
(*与上位机通讯程序*)
ComConveyor70104(ConveyorIO:= ConveyorIO70140_1,CommunicationIO:= ComConveyorIO70104);
ComConveyor70106(ConveyorIO:= ConveyorIO70140,CommunicationIO:= ComConveyorIO70106);(*线体更改*)
ComConveyor70144(ConveyorIO:= ConveyorIO70144,CommunicationIO:= ComConveyorIO70144);
ComConveyor70152(ConveyorIO:= ConveyorIO70152,CommunicationIO:= ComConveyorIO70152);
ComConveyor70146(ConveyorIO:= ConveyorIO70146,CommunicationIO:= ComConveyorIO70146);
ComConveyor70195(ConveyorIO:= ConveyorIO70195,CommunicationIO:= ComConveyorIO70195);
ComConveyor70147(ConveyorIO:= ConveyorIO70147,CommunicationIO:= ComConveyorIO70147);
ComConveyor70196(ConveyorIO:= ConveyorIO70196,CommunicationIO:= ComConveyorIO70196);
ComConveyor70154(ConveyorIO:= ConveyorIO70154,CommunicationIO:= ComConveyorIO70154);
ComConveyor70199(ConveyorIO:= ConveyorIO70199,CommunicationIO:= ComConveyorIO70199);
ComConveyor70155(ConveyorIO:= ConveyorIO70155,CommunicationIO:= ComConveyorIO70155);
ComConveyor701100(ConveyorIO:= ConveyorIO701100,CommunicationIO:= ComConveyorIO701100);
ComConveyor701115(ConveyorIO:= ConveyorIO701115,CommunicationIO:= ComConveyorIO701115);
ComConveyor701114(ConveyorIO:= ConveyorIO701114,CommunicationIO:= ComConveyorIO701114);
ComConveyor70197(ConveyorIO:= ConveyorIO70197,CommunicationIO:= ComConveyorIO70197);
ComConveyor70150(ConveyorIO:= ConveyorIO70150,CommunicationIO:= ComConveyorIO70150);
ComConveyor70151(ConveyorIO:= ConveyorIO70151,CommunicationIO:= ComConveyorIO70151);
ComConveyor70198(ConveyorIO:= ConveyorIO70198,CommunicationIO:= ComConveyorIO70198);
ComConveyor701101(ConveyorIO:= ConveyorIO701101,CommunicationIO:= ComConveyorIO701101);
ComConveyor70158(ConveyorIO:= ConveyorIO70158,CommunicationIO:= ComConveyorIO70158);
ComConveyor701111(ConveyorIO:= ConveyorIO701111,CommunicationIO:= ComConveyorIO701111);
ComConveyor70148(ConveyorIO:= ConveyorIO70148,CommunicationIO:= ComConveyorIO70148);
ComConveyor70156(ConveyorIO:= ConveyorIO70156,CommunicationIO:= ComConveyorIO70156);
ComConveyor701116(ConveyorIO:= ConveyorIO701116,CommunicationIO:= ComConveyorIO701116);
ComConveyor70164(ConveyorIO:= ConveyorIO70164,CommunicationIO:= ComConveyorIO70164);
ComConveyor70174(ConveyorIO:= ConveyorIO70174,CommunicationIO:= ComConveyorIO70174);
ComConveyor70169(ConveyorIO:= ConveyorIO70169,CommunicationIO:= ComConveyorIO70169);
ComConveyor70170(ConveyorIO:= ConveyorIO70170,CommunicationIO:= ComConveyorIO70170);
ComConveyor70160(ConveyorIO:= ConveyorIO70160,CommunicationIO:= ComConveyorIO70160);
ComConveyor70162(ConveyorIO:= ConveyorIO70162,CommunicationIO:= ComConveyorIO70162);
ComConveyor701103(ConveyorIO:= ConveyorIO701103,CommunicationIO:= ComConveyorIO701103);
ComConveyor70163(ConveyorIO:= ConveyorIO70163,CommunicationIO:= ComConveyorIO70163);
ComConveyor701104(ConveyorIO:= ConveyorIO701104,CommunicationIO:= ComConveyorIO701104);
ComConveyor701102(ConveyorIO:= ConveyorIO701102,CommunicationIO:= ComConveyorIO701102);
ComConveyor70159(ConveyorIO:= ConveyorIO70159,CommunicationIO:= ComConveyorIO70159);
ComConveyor701120(ConveyorIO:= ConveyorIO701120,CommunicationIO:= ComConveyorIO701120);
ComConveyor701119(ConveyorIO:= ConveyorIO701119,CommunicationIO:= ComConveyorIO701119);
(*ComConveyor70111(ConveyorIO:= ConveyorIO70111,CommunicationIO:= ComConveyorIO70111);
ComConveyor70112(ConveyorIO:= ConveyorIO70112,CommunicationIO:= ComConveyorIO70112);
ComConveyor701105(ConveyorIO:= ConveyorIO701105,CommunicationIO:= ComConveyorIO701105);
ComConveyor70113(ConveyorIO:= ConveyorIO70113,CommunicationIO:= ComConveyorIO70113);
ComConveyor701106(ConveyorIO:= ConveyorIO701106,CommunicationIO:= ComConveyorIO701106);
ComConveyor70114(ConveyorIO:= ConveyorIO70114,CommunicationIO:= ComConveyorIO70114);
ComConveyor70116(ConveyorIO:= ConveyorIO70116,CommunicationIO:= ComConveyorIO70116);
ComConveyor70119(ConveyorIO:= ConveyorIO70119,CommunicationIO:= ComConveyorIO70119);
ComConveyor70120(ConveyorIO:= ConveyorIO70120,CommunicationIO:= ComConveyorIO70120);
ComConveyor701107(ConveyorIO:= ConveyorIO701107,CommunicationIO:= ComConveyorIO701107);
ComConveyor70121(ConveyorIO:= ConveyorIO70121,CommunicationIO:= ComConveyorIO70121);
ComConveyor701108(ConveyorIO:= ConveyorIO701108,CommunicationIO:= ComConveyorIO701108);
ComConveyor70122(ConveyorIO:= ConveyorIO70122,CommunicationIO:= ComConveyorIO70122);
ComConveyor70124(ConveyorIO:= ConveyorIO70124,CommunicationIO:= ComConveyorIO70124);
ComConveyor70127(ConveyorIO:= ConveyorIO70127,CommunicationIO:= ComConveyorIO70127);
ComConveyor70128(ConveyorIO:= ConveyorIO70128,CommunicationIO:= ComConveyorIO70128);
ComConveyor701109(ConveyorIO:= ConveyorIO701109,CommunicationIO:= ComConveyorIO701109);
ComConveyor70129(ConveyorIO:= ConveyorIO70129,CommunicationIO:= ComConveyorIO70129);
ComConveyor701110(ConveyorIO:= ConveyorIO701110,CommunicationIO:= ComConveyorIO701110);
ComConveyor70184(ConveyorIO:= ConveyorIO70184,CommunicationIO:= ComConveyorIO70184);*)

ComConveyorIO70104.i_iResponsPCPLC:=D2000; 
ComConveyorIO70104.i_iTypeInfoPCPLC:=D2001;
ComConveyorIO70104.i_iReadWriteFlagPCPLC:=D2005; 
ComConveyorIO70104.i_iTaskProcessFlagPCPLC:=D2006; 
ComConveyorIO70104.i_iCommandPCPLC:=D2007; 
ComConveyorIO70104.i_iTaskIDPCPLC:=D2008; 
DMOV(TRUE,D2009,ComConveyorIO70104.i_diDestinationDevicePCPLC); 
ComConveyorIO70104.i_iProductIDPCPLC:=D2011;
D3000:=ComConveyorIO70104.o_iRequestPLCPC; 
D3001:=ComConveyorIO70104.o_iForceInportPLCPC;
D3002:=ComConveyorIO70104.o_iFolderNumberPLCPC;
D3003:=ComConveyorIO70104.o_iEmptyPLCPC;
D3005:=ComConveyorIO70104.o_iReadWriteFlagPLCPC; 
D3006:=ComConveyorIO70104.o_iDeviceStatusPLCPC; 
D3007:=ComConveyorIO70104.o_iTaskIDPLCPC; 
D3008:=ComConveyorIO70104.o_iProductIDPLCPC;

ComConveyorIO70106.i_iTypeInfoPCPLC:=D2031;
ComConveyorIO70106.i_iReadWriteFlagPCPLC:=D2035; 
ComConveyorIO70106.i_iTaskProcessFlagPCPLC:=D2036; 
ComConveyorIO70106.i_iCommandPCPLC:=D2037; 
ComConveyorIO70106.i_iTaskIDPCPLC:=D2038; 
DMOV(TRUE,D2039,ComConveyorIO70106.i_diDestinationDevicePCPLC); 
ComConveyorIO70106.i_iProductIDPCPLC:=D2041;
D3030:=ComConveyorIO70106.o_iRequestPLCPC; 
D3031:=ComConveyorIO70106.o_iForceInportPLCPC;
D3032:=ComConveyorIO70106.o_iFolderNumberPLCPC;
D3033:=ComConveyorIO70106.o_iEmptyPLCPC;
D3035:=ComConveyorIO70106.o_iReadWriteFlagPLCPC; 
D3036:=ComConveyorIO70106.o_iDeviceStatusPLCPC; 
D3037:=ComConveyorIO70106.o_iTaskIDPLCPC; 
D3038:=ComConveyorIO70106.o_iProductIDPLCPC;
ComConveyorIO70144.i_iResponsPCPLC:=D2045; 
ComConveyorIO70144.i_iTypeInfoPCPLC:=D2046;
ComConveyorIO70144.i_iReadWriteFlagPCPLC:=D2050; 
ComConveyorIO70144.i_iTaskProcessFlagPCPLC:=D2051; 
ComConveyorIO70144.i_iCommandPCPLC:=D2052; 
ComConveyorIO70144.i_iTaskIDPCPLC:=D2053; 
DMOV(TRUE,D2054,ComConveyorIO70144.i_diDestinationDevicePCPLC); 
ComConveyorIO70144.i_iProductIDPCPLC:=D2056;
D3045:=ComConveyorIO70144.o_iRequestPLCPC; 
D3046:=ComConveyorIO70144.o_iForceInportPLCPC;
D3047:=ComConveyorIO70144.o_iFolderNumberPLCPC;
D3048:=ComConveyorIO70144.o_iEmptyPLCPC;
D3050:=ComConveyorIO70144.o_iReadWriteFlagPLCPC; 
D3051:=ComConveyorIO70144.o_iDeviceStatusPLCPC; 
D3052:=ComConveyorIO70144.o_iTaskIDPLCPC; 
D3053:=ComConveyorIO70144.o_iProductIDPLCPC;
ComConveyorIO70152.i_iResponsPCPLC:=D2060; 
ComConveyorIO70152.i_iTypeInfoPCPLC:=D2061;
ComConveyorIO70152.i_iReadWriteFlagPCPLC:=D2065; 
ComConveyorIO70152.i_iTaskProcessFlagPCPLC:=D2066; 
ComConveyorIO70152.i_iCommandPCPLC:=D2067; 
ComConveyorIO70152.i_iTaskIDPCPLC:=D2068; 
DMOV(TRUE,D2069,ComConveyorIO70152.i_diDestinationDevicePCPLC); 
ComConveyorIO70152.i_iProductIDPCPLC:=D2071;
D3060:=ComConveyorIO70152.o_iRequestPLCPC; 
D3061:=ComConveyorIO70152.o_iForceInportPLCPC;
D3062:=ComConveyorIO70152.o_iFolderNumberPLCPC;
D3063:=ComConveyorIO70152.o_iEmptyPLCPC;
D3065:=ComConveyorIO70152.o_iReadWriteFlagPLCPC; 
D3066:=ComConveyorIO70152.o_iDeviceStatusPLCPC; 
D3067:=ComConveyorIO70152.o_iTaskIDPLCPC; 
D3068:=ComConveyorIO70152.o_iProductIDPLCPC;
ComConveyorIO70146.i_iResponsPCPLC:=D2075; 
ComConveyorIO70146.i_iTypeInfoPCPLC:=D2076;
ComConveyorIO70146.i_iReadWriteFlagPCPLC:=D2080; 
ComConveyorIO70146.i_iTaskProcessFlagPCPLC:=D2081; 
ComConveyorIO70146.i_iCommandPCPLC:=D2082; 
ComConveyorIO70146.i_iTaskIDPCPLC:=D2083; 
DMOV(TRUE,D2084,ComConveyorIO70146.i_diDestinationDevicePCPLC); 
ComConveyorIO70146.i_iProductIDPCPLC:=D2086;
D3075:=ComConveyorIO70146.o_iRequestPLCPC; 
D3076:=ComConveyorIO70146.o_iForceInportPLCPC;
D3077:=ComConveyorIO70146.o_iFolderNumberPLCPC;
D3078:=ComConveyorIO70146.o_iEmptyPLCPC;
D3080:=ComConveyorIO70146.o_iReadWriteFlagPLCPC; 
D3081:=ComConveyorIO70146.o_iDeviceStatusPLCPC; 
D3082:=ComConveyorIO70146.o_iTaskIDPLCPC; 
D3083:=ComConveyorIO70146.o_iProductIDPLCPC;
ComConveyorIO70195.i_iResponsPCPLC:=D2090; 
ComConveyorIO70195.i_iTypeInfoPCPLC:=D2091;
ComConveyorIO70195.i_iReadWriteFlagPCPLC:=D2095; 
ComConveyorIO70195.i_iTaskProcessFlagPCPLC:=D2096; 
ComConveyorIO70195.i_iCommandPCPLC:=D2097; 
ComConveyorIO70195.i_iTaskIDPCPLC:=D2098; 
DMOV(TRUE,D2099,ComConveyorIO70195.i_diDestinationDevicePCPLC); 
ComConveyorIO70195.i_iProductIDPCPLC:=D2101;
D3090:=ComConveyorIO70195.o_iRequestPLCPC; 
D3091:=ComConveyorIO70195.o_iForceInportPLCPC;
D3092:=ComConveyorIO70195.o_iFolderNumberPLCPC;
D3093:=ComConveyorIO70195.o_iEmptyPLCPC;
D3095:=ComConveyorIO70195.o_iReadWriteFlagPLCPC; 
D3096:=ComConveyorIO70195.o_iDeviceStatusPLCPC; 
D3097:=ComConveyorIO70195.o_iTaskIDPLCPC; 
D3098:=ComConveyorIO70195.o_iProductIDPLCPC;
ComConveyorIO70147.i_iResponsPCPLC:=D2105; 
ComConveyorIO70147.i_iTypeInfoPCPLC:=D2106;
ComConveyorIO70147.i_iReadWriteFlagPCPLC:=D2110; 
ComConveyorIO70147.i_iTaskProcessFlagPCPLC:=D2111; 
ComConveyorIO70147.i_iCommandPCPLC:=D2112; 
ComConveyorIO70147.i_iTaskIDPCPLC:=D2113; 
DMOV(TRUE,D2114,ComConveyorIO70147.i_diDestinationDevicePCPLC); 
ComConveyorIO70147.i_iProductIDPCPLC:=D2116;
D3105:=ComConveyorIO70147.o_iRequestPLCPC; 
D3106:=ComConveyorIO70147.o_iForceInportPLCPC;
D3107:=ComConveyorIO70147.o_iFolderNumberPLCPC;
D3108:=ComConveyorIO70147.o_iEmptyPLCPC;
D3110:=ComConveyorIO70147.o_iReadWriteFlagPLCPC; 
D3111:=ComConveyorIO70147.o_iDeviceStatusPLCPC; 
D3112:=ComConveyorIO70147.o_iTaskIDPLCPC; 
D3113:=ComConveyorIO70147.o_iProductIDPLCPC;
ComConveyorIO70196.i_iResponsPCPLC:=D2120; 
ComConveyorIO70196.i_iTypeInfoPCPLC:=D2121;
ComConveyorIO70196.i_iReadWriteFlagPCPLC:=D2125; 
ComConveyorIO70196.i_iTaskProcessFlagPCPLC:=D2126; 
ComConveyorIO70196.i_iCommandPCPLC:=D2127; 
ComConveyorIO70196.i_iTaskIDPCPLC:=D2128; 
DMOV(TRUE,D2129,ComConveyorIO70196.i_diDestinationDevicePCPLC); 
ComConveyorIO70196.i_iProductIDPCPLC:=D2131;	
D3120:=ComConveyorIO70196.o_iRequestPLCPC; 
D3121:=ComConveyorIO70196.o_iForceInportPLCPC;
D3122:=ComConveyorIO70196.o_iFolderNumberPLCPC;
D3123:=ComConveyorIO70196.o_iEmptyPLCPC;
D3125:=ComConveyorIO70196.o_iReadWriteFlagPLCPC; 
D3126:=ComConveyorIO70196.o_iDeviceStatusPLCPC; 
D3127:=ComConveyorIO70196.o_iTaskIDPLCPC; 
D3128:=ComConveyorIO70196.o_iProductIDPLCPC;
ComConveyorIO70154.i_iResponsPCPLC:=D2135; 
ComConveyorIO70154.i_iTypeInfoPCPLC:=D2136;
ComConveyorIO70154.i_iReadWriteFlagPCPLC:=D2140; 
ComConveyorIO70154.i_iTaskProcessFlagPCPLC:=D2141; 
ComConveyorIO70154.i_iCommandPCPLC:=D2142; 
ComConveyorIO70154.i_iTaskIDPCPLC:=D2143; 
DMOV(TRUE,D2144,ComConveyorIO70154.i_diDestinationDevicePCPLC); 
ComConveyorIO70154.i_iProductIDPCPLC:=D2146;
D3135:=ComConveyorIO70154.o_iRequestPLCPC; 
D3136:=ComConveyorIO70154.o_iForceInportPLCPC;
D3137:=ComConveyorIO70154.o_iFolderNumberPLCPC;
D3138:=ComConveyorIO70154.o_iEmptyPLCPC;
D3140:=ComConveyorIO70154.o_iReadWriteFlagPLCPC; 
D3141:=ComConveyorIO70154.o_iDeviceStatusPLCPC; 
D3142:=ComConveyorIO70154.o_iTaskIDPLCPC; 
D3143:=ComConveyorIO70154.o_iProductIDPLCPC;
ComConveyorIO70199.i_iResponsPCPLC:=D2150; 
ComConveyorIO70199.i_iTypeInfoPCPLC:=D2151;
ComConveyorIO70199.i_iReadWriteFlagPCPLC:=D2155; 
ComConveyorIO70199.i_iTaskProcessFlagPCPLC:=D2156; 
ComConveyorIO70199.i_iCommandPCPLC:=D2157; 
ComConveyorIO70199.i_iTaskIDPCPLC:=D2158; 
DMOV(TRUE,D2159,ComConveyorIO70199.i_diDestinationDevicePCPLC); 
ComConveyorIO70199.i_iProductIDPCPLC:=D2161;
D3150:=ComConveyorIO70199.o_iRequestPLCPC; 
D3151:=ComConveyorIO70199.o_iForceInportPLCPC;
D3152:=ComConveyorIO70199.o_iFolderNumberPLCPC;
D3153:=ComConveyorIO70199.o_iEmptyPLCPC;
D3155:=ComConveyorIO70199.o_iReadWriteFlagPLCPC; 
D3156:=ComConveyorIO70199.o_iDeviceStatusPLCPC; 
D3157:=ComConveyorIO70199.o_iTaskIDPLCPC; 
D3158:=ComConveyorIO70199.o_iProductIDPLCPC;
ComConveyorIO70155.i_iResponsPCPLC:=D2165; 
ComConveyorIO70155.i_iTypeInfoPCPLC:=D2166;
ComConveyorIO70155.i_iReadWriteFlagPCPLC:=D2170; 
ComConveyorIO70155.i_iTaskProcessFlagPCPLC:=D2171; 
ComConveyorIO70155.i_iCommandPCPLC:=D2172; 
ComConveyorIO70155.i_iTaskIDPCPLC:=D2173; 
DMOV(TRUE,D2174,ComConveyorIO70155.i_diDestinationDevicePCPLC); 
ComConveyorIO70155.i_iProductIDPCPLC:=D2176;	
D3165:=ComConveyorIO70155.o_iRequestPLCPC; 
D3166:=ComConveyorIO70155.o_iForceInportPLCPC;
D3167:=ComConveyorIO70155.o_iFolderNumberPLCPC;
D3168:=ComConveyorIO70155.o_iEmptyPLCPC;
D3170:=ComConveyorIO70155.o_iReadWriteFlagPLCPC; 
D3171:=ComConveyorIO70155.o_iDeviceStatusPLCPC; 
D3172:=ComConveyorIO70155.o_iTaskIDPLCPC; 
D3173:=ComConveyorIO70155.o_iProductIDPLCPC;
ComConveyorIO701100.i_iResponsPCPLC:=D2180; 
ComConveyorIO701100.i_iTypeInfoPCPLC:=D2181;
ComConveyorIO701100.i_iReadWriteFlagPCPLC:=D2185; 
ComConveyorIO701100.i_iTaskProcessFlagPCPLC:=D2186; 
ComConveyorIO701100.i_iCommandPCPLC:=D2187; 
ComConveyorIO701100.i_iTaskIDPCPLC:=D2188; 
DMOV(TRUE,D2189,ComConveyorIO701100.i_diDestinationDevicePCPLC); 
ComConveyorIO701100.i_iProductIDPCPLC:=D2191;
D3180:=ComConveyorIO701100.o_iRequestPLCPC; 
D3181:=ComConveyorIO701100.o_iForceInportPLCPC;
D3182:=ComConveyorIO701100.o_iFolderNumberPLCPC;
D3183:=ComConveyorIO701100.o_iEmptyPLCPC;
D3185:=ComConveyorIO701100.o_iReadWriteFlagPLCPC; 
D3186:=ComConveyorIO701100.o_iDeviceStatusPLCPC; 
D3187:=ComConveyorIO701100.o_iTaskIDPLCPC; 
D3188:=ComConveyorIO701100.o_iProductIDPLCPC;
ComConveyorIO701115.i_iResponsPCPLC:=D2195; 
ComConveyorIO701115.i_iTypeInfoPCPLC:=D2196;
ComConveyorIO701115.i_iReadWriteFlagPCPLC:=D2200; 
ComConveyorIO701115.i_iTaskProcessFlagPCPLC:=D2201; 
ComConveyorIO701115.i_iCommandPCPLC:=D2202; 
ComConveyorIO701115.i_iTaskIDPCPLC:=D2203; 
DMOV(TRUE,D2204,ComConveyorIO701115.i_diDestinationDevicePCPLC); 
ComConveyorIO701115.i_iProductIDPCPLC:=D2206;
D3195:=ComConveyorIO701115.o_iRequestPLCPC; 
D3196:=ComConveyorIO701115.o_iForceInportPLCPC;
D3197:=ComConveyorIO701115.o_iFolderNumberPLCPC;
D3198:=ComConveyorIO701115.o_iEmptyPLCPC;
D3200:=ComConveyorIO701115.o_iReadWriteFlagPLCPC; 
D3201:=ComConveyorIO701115.o_iDeviceStatusPLCPC; 
D3202:=ComConveyorIO701115.o_iTaskIDPLCPC; 
D3203:=ComConveyorIO701115.o_iProductIDPLCPC;
ComConveyorIO701115.i_xExportConveyor:=1;
ComConveyorIO701115.i_xExtraCondition:=ConveyorIO701114.xEmpty AND NOT ConveyorIO701114.xCWPresent AND NOT ConveyorIO701115.xCWPresent;

(*ComConveyorIO701114.i_iResponsPCPLC:=D2210; 
ComConveyorIO701114.i_iTypeInfoPCPLC:=D2211;
ComConveyorIO701114.i_iReadWriteFlagPCPLC:=D2215; 
ComConveyorIO701114.i_iTaskProcessFlagPCPLC:=D2216; 
ComConveyorIO701114.i_iCommandPCPLC:=D2217; 
ComConveyorIO701114.i_iTaskIDPCPLC:=D2218; 
DMOV(TRUE,D2219,ComConveyorIO701114.i_diDestinationDevicePCPLC); 
ComConveyorIO701114.i_iProductIDPCPLC:=D2221;
D3210:=ComConveyorIO701114.o_iRequestPLCPC; 
D3211:=ComConveyorIO701114.o_iForceInportPLCPC;
D3212:=ComConveyorIO701114.o_iFolderNumberPLCPC;
D3213:=ComConveyorIO701114.o_iEmptyPLCPC;
D3215:=ComConveyorIO701114.o_iReadWriteFlagPLCPC; 
D3216:=ComConveyorIO701114.o_iDeviceStatusPLCPC; 
D3217:=ComConveyorIO701114.o_iTaskIDPLCPC; 
D3218:=ComConveyorIO701114.o_iProductIDPLCPC;
ComConveyorIO701114.i_xExportConveyor:=1;*)

ComConveyorIO70197.i_iResponsPCPLC:=D2225; 
ComConveyorIO70197.i_iTypeInfoPCPLC:=D2226;
ComConveyorIO70197.i_iReadWriteFlagPCPLC:=D2230; 
ComConveyorIO70197.i_iTaskProcessFlagPCPLC:=D2231; 
ComConveyorIO70197.i_iCommandPCPLC:=D2232; 
ComConveyorIO70197.i_iTaskIDPCPLC:=D2233; 
DMOV(TRUE,D2234,ComConveyorIO70197.i_diDestinationDevicePCPLC); 
ComConveyorIO70197.i_iProductIDPCPLC:=D2236;
D3225:=ComConveyorIO70197.o_iRequestPLCPC; 
D3226:=ComConveyorIO70197.o_iForceInportPLCPC;
D3227:=ComConveyorIO70197.o_iFolderNumberPLCPC;
D3228:=ComConveyorIO70197.o_iEmptyPLCPC;
D3230:=ComConveyorIO70197.o_iReadWriteFlagPLCPC; 
D3231:=ComConveyorIO70197.o_iDeviceStatusPLCPC; 
D3232:=ComConveyorIO70197.o_iTaskIDPLCPC; 
D3233:=ComConveyorIO70197.o_iProductIDPLCPC;
ComConveyorIO70197.i_xExportConveyor:=1;
ComConveyorIO70197.i_xExtraCondition:=ConveyorIO70150.xEmpty AND NOT ConveyorIO70150.xCWPresent AND NOT ConveyorIO70197.xCWPresent;
(*
ComConveyorIO70150.i_iResponsPCPLC:=D2240; 
ComConveyorIO70150.i_iTypeInfoPCPLC:=D2241;
ComConveyorIO70150.i_iReadWriteFlagPCPLC:=D2245; 
ComConveyorIO70150.i_iTaskProcessFlagPCPLC:=D2246; 
ComConveyorIO70150.i_iCommandPCPLC:=D2247; 
ComConveyorIO70150.i_iTaskIDPCPLC:=D2248; 
DMOV(TRUE,D2249,ComConveyorIO70150.i_diDestinationDevicePCPLC); 
ComConveyorIO70150.i_iProductIDPCPLC:=D2251;
D3240:=ComConveyorIO70150.o_iRequestPLCPC; 
D3241:=ComConveyorIO70150.o_iForceInportPLCPC;
D3242:=ComConveyorIO70150.o_iFolderNumberPLCPC;
D3243:=ComConveyorIO70150.o_iEmptyPLCPC;
D3245:=ComConveyorIO70150.o_iReadWriteFlagPLCPC; 
D3246:=ComConveyorIO70150.o_iDeviceStatusPLCPC; 
D3247:=ComConveyorIO70150.o_iTaskIDPLCPC; 
D3248:=ComConveyorIO70150.o_iProductIDPLCPC;
ComConveyorIO70150.i_xExportConveyor:=1;*)

ComConveyorIO70151.i_iResponsPCPLC:=D2255; 
ComConveyorIO70151.i_iTypeInfoPCPLC:=D2256;
ComConveyorIO70151.i_iReadWriteFlagPCPLC:=D2260; 
ComConveyorIO70151.i_iTaskProcessFlagPCPLC:=D2261; 
ComConveyorIO70151.i_iCommandPCPLC:=D2262; 
ComConveyorIO70151.i_iTaskIDPCPLC:=D2263; 
DMOV(TRUE,D2264,ComConveyorIO70151.i_diDestinationDevicePCPLC); 
ComConveyorIO70151.i_iProductIDPCPLC:=D2266;
D3255:=ComConveyorIO70151.o_iRequestPLCPC; 
D3256:=ComConveyorIO70151.o_iForceInportPLCPC;
D3257:=ComConveyorIO70151.o_iFolderNumberPLCPC;
D3258:=ComConveyorIO70151.o_iEmptyPLCPC;
D3260:=ComConveyorIO70151.o_iReadWriteFlagPLCPC; 
D3261:=ComConveyorIO70151.o_iDeviceStatusPLCPC; 
D3262:=ComConveyorIO70151.o_iTaskIDPLCPC; 
D3263:=ComConveyorIO70151.o_iProductIDPLCPC;
ComConveyorIO70151.i_xExportConveyor:=1;
ComConveyorIO70151.i_xExtraCondition:=ConveyorIO70198.xEmpty AND NOT ConveyorIO70198.xCWPresent AND NOT ConveyorIO70151.xCWPresent;
(*
ComConveyorIO70198.i_iResponsPCPLC:=D2270; 
ComConveyorIO70198.i_iTypeInfoPCPLC:=D2271;
ComConveyorIO70198.i_iReadWriteFlagPCPLC:=D2275; 
ComConveyorIO70198.i_iTaskProcessFlagPCPLC:=D2276; 
ComConveyorIO70198.i_iCommandPCPLC:=D2277; 
ComConveyorIO70198.i_iTaskIDPCPLC:=D2278; 
DMOV(TRUE,D2279,ComConveyorIO70198.i_diDestinationDevicePCPLC); 
ComConveyorIO70198.i_iProductIDPCPLC:=D2281;
D3270:=ComConveyorIO70198.o_iRequestPLCPC; 
D3271:=ComConveyorIO70198.o_iForceInportPLCPC;
D3272:=ComConveyorIO70198.o_iFolderNumberPLCPC;
D3273:=ComConveyorIO70198.o_iEmptyPLCPC;
D3275:=ComConveyorIO70198.o_iReadWriteFlagPLCPC; 
D3276:=ComConveyorIO70198.o_iDeviceStatusPLCPC; 
D3277:=ComConveyorIO70198.o_iTaskIDPLCPC; 
D3278:=ComConveyorIO70198.o_iProductIDPLCPC;
ComConveyorIO70198.i_xExportConveyor:=1;*)

ComConveyorIO701101.i_iResponsPCPLC:=D2285; 
ComConveyorIO701101.i_iTypeInfoPCPLC:=D2286;
ComConveyorIO701101.i_iReadWriteFlagPCPLC:=D2290; 
ComConveyorIO701101.i_iTaskProcessFlagPCPLC:=D2291; 
ComConveyorIO701101.i_iCommandPCPLC:=D2292; 
ComConveyorIO701101.i_iTaskIDPCPLC:=D2293; 
DMOV(TRUE,D2294,ComConveyorIO701101.i_diDestinationDevicePCPLC); 
ComConveyorIO701101.i_iProductIDPCPLC:=D2296;
D3285:=ComConveyorIO701101.o_iRequestPLCPC; 
D3286:=ComConveyorIO701101.o_iForceInportPLCPC;
D3287:=ComConveyorIO701101.o_iFolderNumberPLCPC;
D3288:=ComConveyorIO701101.o_iEmptyPLCPC;
D3290:=ComConveyorIO701101.o_iReadWriteFlagPLCPC; 
D3291:=ComConveyorIO701101.o_iDeviceStatusPLCPC; 
D3292:=ComConveyorIO701101.o_iTaskIDPLCPC; 
D3293:=ComConveyorIO701101.o_iProductIDPLCPC;
ComConveyorIO701101.i_xExportConveyor:=1;
ComConveyorIO701101.i_xExtraCondition:=ConveyorIO70158.xEmpty AND NOT ConveyorIO70158.xCWPresent AND NOT ConveyorIO701101.xCWPresent;
(*
ComConveyorIO70158.i_iResponsPCPLC:=D2300; 
ComConveyorIO70158.i_iTypeInfoPCPLC:=D2301;
ComConveyorIO70158.i_iReadWriteFlagPCPLC:=D2305; 
ComConveyorIO70158.i_iTaskProcessFlagPCPLC:=D2306; 
ComConveyorIO70158.i_iCommandPCPLC:=D2307; 
ComConveyorIO70158.i_iTaskIDPCPLC:=D2308; 
DMOV(TRUE,D2309,ComConveyorIO70158.i_diDestinationDevicePCPLC); 
ComConveyorIO70158.i_iProductIDPCPLC:=D2311;
D3300:=ComConveyorIO70158.o_iRequestPLCPC; 
D3301:=ComConveyorIO70158.o_iForceInportPLCPC;
D3302:=ComConveyorIO70158.o_iFolderNumberPLCPC;
D3303:=ComConveyorIO70158.o_iEmptyPLCPC;
D3305:=ComConveyorIO70158.o_iReadWriteFlagPLCPC; 
D3306:=ComConveyorIO70158.o_iDeviceStatusPLCPC; 
D3307:=ComConveyorIO70158.o_iTaskIDPLCPC; 
D3308:=ComConveyorIO70158.o_iProductIDPLCPC;
ComConveyorIO70158.i_xExportConveyor:=1;*)

ComConveyorIO701111.i_iResponsPCPLC:=D2315; 
ComConveyorIO701111.i_iTypeInfoPCPLC:=D2316;
ComConveyorIO701111.i_iReadWriteFlagPCPLC:=D2320; 
ComConveyorIO701111.i_iTaskProcessFlagPCPLC:=D2321; 
ComConveyorIO701111.i_iCommandPCPLC:=D2322; 
ComConveyorIO701111.i_iTaskIDPCPLC:=D2323; 
DMOV(TRUE,D2324,ComConveyorIO701111.i_diDestinationDevicePCPLC); 
ComConveyorIO701111.i_iProductIDPCPLC:=D2326;
D3315:=ComConveyorIO701111.o_iRequestPLCPC; 
D3316:=ComConveyorIO701111.o_iForceInportPLCPC;
D3317:=ComConveyorIO701111.o_iFolderNumberPLCPC;
D3318:=ComConveyorIO701111.o_iEmptyPLCPC;
D3320:=ComConveyorIO701111.o_iReadWriteFlagPLCPC; 
D3321:=ComConveyorIO701111.o_iDeviceStatusPLCPC; 
D3322:=ComConveyorIO701111.o_iTaskIDPLCPC; 
D3323:=ComConveyorIO701111.o_iProductIDPLCPC;
ComConveyorIO70148.i_iResponsPCPLC:=D2330; 
ComConveyorIO70148.i_iTypeInfoPCPLC:=D2331;
ComConveyorIO70148.i_iReadWriteFlagPCPLC:=D2335; 
ComConveyorIO70148.i_iTaskProcessFlagPCPLC:=D2336; 
ComConveyorIO70148.i_iCommandPCPLC:=D2337; 
ComConveyorIO70148.i_iTaskIDPCPLC:=D2338; 
DMOV(TRUE,D2339,ComConveyorIO70148.i_diDestinationDevicePCPLC); 
ComConveyorIO70148.i_iProductIDPCPLC:=D2341;
D3330:=ComConveyorIO70148.o_iRequestPLCPC; 
D3331:=ComConveyorIO70148.o_iForceInportPLCPC;
D3332:=ComConveyorIO70148.o_iFolderNumberPLCPC;
D3333:=ComConveyorIO70148.o_iEmptyPLCPC;
D3335:=ComConveyorIO70148.o_iReadWriteFlagPLCPC; 
D3336:=ComConveyorIO70148.o_iDeviceStatusPLCPC; 
D3337:=ComConveyorIO70148.o_iTaskIDPLCPC; 
D3338:=ComConveyorIO70148.o_iProductIDPLCPC;
ComConveyorIO70156.i_iResponsPCPLC:=D2345; 
ComConveyorIO70156.i_iTypeInfoPCPLC:=D2346;
ComConveyorIO70156.i_iReadWriteFlagPCPLC:=D2350; 
ComConveyorIO70156.i_iTaskProcessFlagPCPLC:=D2351; 
ComConveyorIO70156.i_iCommandPCPLC:=D2352; 
ComConveyorIO70156.i_iTaskIDPCPLC:=D2353; 
DMOV(TRUE,D2354,ComConveyorIO70156.i_diDestinationDevicePCPLC); 
ComConveyorIO70156.i_iProductIDPCPLC:=D2356;
D3345:=ComConveyorIO70156.o_iRequestPLCPC; 
D3346:=ComConveyorIO70156.o_iForceInportPLCPC;
D3347:=ComConveyorIO70156.o_iFolderNumberPLCPC;
D3348:=ComConveyorIO70156.o_iEmptyPLCPC;
D3350:=ComConveyorIO70156.o_iReadWriteFlagPLCPC; 
D3351:=ComConveyorIO70156.o_iDeviceStatusPLCPC; 
D3352:=ComConveyorIO70156.o_iTaskIDPLCPC; 
D3353:=ComConveyorIO70156.o_iProductIDPLCPC;
ComConveyorIO701116.i_iResponsPCPLC:=D2360; 
ComConveyorIO701116.i_iTypeInfoPCPLC:=D2361;
ComConveyorIO701116.i_iReadWriteFlagPCPLC:=D2365; 
ComConveyorIO701116.i_iTaskProcessFlagPCPLC:=D2366; 
ComConveyorIO701116.i_iCommandPCPLC:=D2367; 
ComConveyorIO701116.i_iTaskIDPCPLC:=D2368; 
DMOV(TRUE,D2369,ComConveyorIO701116.i_diDestinationDevicePCPLC); 
ComConveyorIO701116.i_iProductIDPCPLC:=D2371;
D3360:=ComConveyorIO701116.o_iRequestPLCPC; 
D3361:=ComConveyorIO701116.o_iForceInportPLCPC;
D3362:=ComConveyorIO701116.o_iFolderNumberPLCPC;
D3363:=ComConveyorIO701116.o_iEmptyPLCPC;
D3365:=ComConveyorIO701116.o_iReadWriteFlagPLCPC; 
D3366:=ComConveyorIO701116.o_iDeviceStatusPLCPC; 
D3367:=ComConveyorIO701116.o_iTaskIDPLCPC; 
D3368:=ComConveyorIO701116.o_iProductIDPLCPC;
ComConveyorIO70164.i_iResponsPCPLC:=D2375; 
ComConveyorIO70164.i_iTypeInfoPCPLC:=D2376;
ComConveyorIO70164.i_iReadWriteFlagPCPLC:=D2380; 
ComConveyorIO70164.i_iTaskProcessFlagPCPLC:=D2381; 
ComConveyorIO70164.i_iCommandPCPLC:=D2382; 
ComConveyorIO70164.i_iTaskIDPCPLC:=D2383; 
DMOV(TRUE,D2384,ComConveyorIO70164.i_diDestinationDevicePCPLC); 
ComConveyorIO70164.i_iProductIDPCPLC:=D2386;
D3375:=ComConveyorIO70164.o_iRequestPLCPC; 
D3376:=ComConveyorIO70164.o_iForceInportPLCPC;
D3377:=ComConveyorIO70164.o_iFolderNumberPLCPC;
D3378:=ComConveyorIO70164.o_iEmptyPLCPC;
D3380:=ComConveyorIO70164.o_iReadWriteFlagPLCPC; 
D3381:=ComConveyorIO70164.o_iDeviceStatusPLCPC; 
D3382:=ComConveyorIO70164.o_iTaskIDPLCPC; 
D3383:=ComConveyorIO70164.o_iProductIDPLCPC;
ComConveyorIO70174.i_iResponsPCPLC:=D2390; 
ComConveyorIO70174.i_iTypeInfoPCPLC:=D2391;
ComConveyorIO70174.i_iReadWriteFlagPCPLC:=D2395; 
ComConveyorIO70174.i_iTaskProcessFlagPCPLC:=D2396; 
ComConveyorIO70174.i_iCommandPCPLC:=D2397; 
ComConveyorIO70174.i_iTaskIDPCPLC:=D2398; 
DMOV(TRUE,D2399,ComConveyorIO70174.i_diDestinationDevicePCPLC); 
ComConveyorIO70174.i_iProductIDPCPLC:=D2401;
D3390:=ComConveyorIO70174.o_iRequestPLCPC; 
D3391:=ComConveyorIO70174.o_iForceInportPLCPC;
D3392:=ComConveyorIO70174.o_iFolderNumberPLCPC;
D3393:=ComConveyorIO70174.o_iEmptyPLCPC;
D3395:=ComConveyorIO70174.o_iReadWriteFlagPLCPC; 
D3396:=ComConveyorIO70174.o_iDeviceStatusPLCPC; 
D3397:=ComConveyorIO70174.o_iTaskIDPLCPC; 
D3398:=ComConveyorIO70174.o_iProductIDPLCPC;
ComConveyorIO70169.i_iResponsPCPLC:=D2405; 
ComConveyorIO70169.i_iTypeInfoPCPLC:=D2406;
ComConveyorIO70169.i_iReadWriteFlagPCPLC:=D2410; 
ComConveyorIO70169.i_iTaskProcessFlagPCPLC:=D2411; 
ComConveyorIO70169.i_iCommandPCPLC:=D2412; 
ComConveyorIO70169.i_iTaskIDPCPLC:=D2413; 
DMOV(TRUE,D2414,ComConveyorIO70169.i_diDestinationDevicePCPLC); 
ComConveyorIO70169.i_iProductIDPCPLC:=D2416;
D3405:=ComConveyorIO70169.o_iRequestPLCPC; 
D3406:=ComConveyorIO70169.o_iForceInportPLCPC;
D3407:=ComConveyorIO70169.o_iFolderNumberPLCPC;
D3408:=ComConveyorIO70169.o_iEmptyPLCPC;
D3410:=ComConveyorIO70169.o_iReadWriteFlagPLCPC; 
D3411:=ComConveyorIO70169.o_iDeviceStatusPLCPC; 
D3412:=ComConveyorIO70169.o_iTaskIDPLCPC; 
D3413:=ComConveyorIO70169.o_iProductIDPLCPC;
ComConveyorIO70170.i_iTypeInfoPCPLC:=D2436;
ComConveyorIO70170.i_iReadWriteFlagPCPLC:=D2440; 
ComConveyorIO70170.i_iTaskProcessFlagPCPLC:=D2441; 
ComConveyorIO70170.i_iCommandPCPLC:=D2442; 
ComConveyorIO70170.i_iTaskIDPCPLC:=D2443; 
DMOV(TRUE,D2444,ComConveyorIO70170.i_diDestinationDevicePCPLC); 
ComConveyorIO70170.i_iProductIDPCPLC:=D2446;
D3435:=ComConveyorIO70170.o_iRequestPLCPC; 
D3436:=ComConveyorIO70170.o_iForceInportPLCPC;
D3437:=ComConveyorIO70170.o_iFolderNumberPLCPC;
D3438:=ComConveyorIO70170.o_iEmptyPLCPC;
D3440:=ComConveyorIO70170.o_iReadWriteFlagPLCPC; 
D3441:=ComConveyorIO70170.o_iDeviceStatusPLCPC; 
D3442:=ComConveyorIO70170.o_iTaskIDPLCPC; 
D3443:=ComConveyorIO70170.o_iProductIDPLCPC;
ComConveyorIO70160.i_iResponsPCPLC:=D2450; 
ComConveyorIO70160.i_iTypeInfoPCPLC:=D2451;
ComConveyorIO70160.i_iReadWriteFlagPCPLC:=D2455; 
ComConveyorIO70160.i_iTaskProcessFlagPCPLC:=D2456; 
ComConveyorIO70160.i_iCommandPCPLC:=D2457; 
ComConveyorIO70160.i_iTaskIDPCPLC:=D2458; 
DMOV(TRUE,D2459,ComConveyorIO70160.i_diDestinationDevicePCPLC); 
ComConveyorIO70160.i_iProductIDPCPLC:=D2461;
D3450:=ComConveyorIO70160.o_iRequestPLCPC; 
D3451:=ComConveyorIO70160.o_iForceInportPLCPC;
D3452:=ComConveyorIO70160.o_iFolderNumberPLCPC;
D3453:=ComConveyorIO70160.o_iEmptyPLCPC;
D3455:=ComConveyorIO70160.o_iReadWriteFlagPLCPC; 
D3456:=ComConveyorIO70160.o_iDeviceStatusPLCPC; 
D3457:=ComConveyorIO70160.o_iTaskIDPLCPC; 
D3458:=ComConveyorIO70160.o_iProductIDPLCPC;
ComConveyorIO70162.i_iResponsPCPLC:=D2465; 
ComConveyorIO70162.i_iTypeInfoPCPLC:=D2466;
ComConveyorIO70162.i_iReadWriteFlagPCPLC:=D2470; 
ComConveyorIO70162.i_iTaskProcessFlagPCPLC:=D2471; 
ComConveyorIO70162.i_iCommandPCPLC:=D2472; 
ComConveyorIO70162.i_iTaskIDPCPLC:=D2473; 
DMOV(TRUE,D2474,ComConveyorIO70162.i_diDestinationDevicePCPLC); 
ComConveyorIO70162.i_iProductIDPCPLC:=D2476;
D3465:=ComConveyorIO70162.o_iRequestPLCPC; 
D3466:=ComConveyorIO70162.o_iForceInportPLCPC;
D3467:=ComConveyorIO70162.o_iFolderNumberPLCPC;
D3468:=ComConveyorIO70162.o_iEmptyPLCPC;
D3470:=ComConveyorIO70162.o_iReadWriteFlagPLCPC; 
D3471:=ComConveyorIO70162.o_iDeviceStatusPLCPC; 
D3472:=ComConveyorIO70162.o_iTaskIDPLCPC; 
D3473:=ComConveyorIO70162.o_iProductIDPLCPC;
ComConveyorIO701103.i_iResponsPCPLC:=D2480; 
ComConveyorIO701103.i_iTypeInfoPCPLC:=D2481;
ComConveyorIO701103.i_iReadWriteFlagPCPLC:=D2485; 
ComConveyorIO701103.i_iTaskProcessFlagPCPLC:=D2486; 
ComConveyorIO701103.i_iCommandPCPLC:=D2487; 
ComConveyorIO701103.i_iTaskIDPCPLC:=D2488; 
DMOV(TRUE,D2489,ComConveyorIO701103.i_diDestinationDevicePCPLC); 
ComConveyorIO701103.i_iProductIDPCPLC:=D2491;
D3480:=ComConveyorIO701103.o_iRequestPLCPC; 
D3481:=ComConveyorIO701103.o_iForceInportPLCPC;
D3482:=ComConveyorIO701103.o_iFolderNumberPLCPC;
D3483:=ComConveyorIO701103.o_iEmptyPLCPC;
D3485:=ComConveyorIO701103.o_iReadWriteFlagPLCPC; 
D3486:=ComConveyorIO701103.o_iDeviceStatusPLCPC; 
D3487:=ComConveyorIO701103.o_iTaskIDPLCPC; 
D3488:=ComConveyorIO701103.o_iProductIDPLCPC;
ComConveyorIO70163.i_iResponsPCPLC:=D2495; 
ComConveyorIO70163.i_iTypeInfoPCPLC:=D2496;
ComConveyorIO70163.i_iReadWriteFlagPCPLC:=D2500; 
ComConveyorIO70163.i_iTaskProcessFlagPCPLC:=D2501; 
ComConveyorIO70163.i_iCommandPCPLC:=D2502; 
ComConveyorIO70163.i_iTaskIDPCPLC:=D2503; 
DMOV(TRUE,D2504,ComConveyorIO70163.i_diDestinationDevicePCPLC); 
ComConveyorIO70163.i_iProductIDPCPLC:=D2506;
D3495:=ComConveyorIO70163.o_iRequestPLCPC; 
D3496:=ComConveyorIO70163.o_iForceInportPLCPC;
D3497:=ComConveyorIO70163.o_iFolderNumberPLCPC;
D3498:=ComConveyorIO70163.o_iEmptyPLCPC;
D3500:=ComConveyorIO70163.o_iReadWriteFlagPLCPC; 
D3501:=ComConveyorIO70163.o_iDeviceStatusPLCPC; 
D3502:=ComConveyorIO70163.o_iTaskIDPLCPC; 
D3503:=ComConveyorIO70163.o_iProductIDPLCPC;
ComConveyorIO701104.i_iResponsPCPLC:=D2510; 
ComConveyorIO701104.i_iTypeInfoPCPLC:=D2511;
ComConveyorIO701104.i_iReadWriteFlagPCPLC:=D2515; 
ComConveyorIO701104.i_iTaskProcessFlagPCPLC:=D2516; 
ComConveyorIO701104.i_iCommandPCPLC:=D2517; 
ComConveyorIO701104.i_iTaskIDPCPLC:=D2518; 
DMOV(TRUE,D2519,ComConveyorIO701104.i_diDestinationDevicePCPLC); 
ComConveyorIO701104.i_iProductIDPCPLC:=D2521;
D3510:=ComConveyorIO701104.o_iRequestPLCPC; 
D3511:=ComConveyorIO701104.o_iForceInportPLCPC;
D3512:=ComConveyorIO701104.o_iFolderNumberPLCPC;
D3513:=ComConveyorIO701104.o_iEmptyPLCPC;
D3515:=ComConveyorIO701104.o_iReadWriteFlagPLCPC; 
D3516:=ComConveyorIO701104.o_iDeviceStatusPLCPC; 
D3517:=ComConveyorIO701104.o_iTaskIDPLCPC; 
D3518:=ComConveyorIO701104.o_iProductIDPLCPC;

ComConveyorIO701102.i_iResponsPCPLC:=D2525; 
ComConveyorIO701102.i_iTypeInfoPCPLC:=D2526;
ComConveyorIO701102.i_iReadWriteFlagPCPLC:=D2530; 
ComConveyorIO701102.i_iTaskProcessFlagPCPLC:=D2531; 
ComConveyorIO701102.i_iCommandPCPLC:=D2532; 
ComConveyorIO701102.i_iTaskIDPCPLC:=D2533; 
DMOV(TRUE,D2534,ComConveyorIO701102.i_diDestinationDevicePCPLC); 
ComConveyorIO701102.i_iProductIDPCPLC:=D2536;
D3525:=ComConveyorIO701102.o_iRequestPLCPC; 
D3526:=ComConveyorIO701102.o_iForceInportPLCPC;
D3527:=ComConveyorIO701102.o_iFolderNumberPLCPC;
D3528:=ComConveyorIO701102.o_iEmptyPLCPC;
D3530:=ComConveyorIO701102.o_iReadWriteFlagPLCPC; 
D3531:=ComConveyorIO701102.o_iDeviceStatusPLCPC; 
D3532:=ComConveyorIO701102.o_iTaskIDPLCPC; 
D3533:=ComConveyorIO701102.o_iProductIDPLCPC;
ComConveyorIO701102.i_xExportConveyor:=1;
ComConveyorIO701102.i_xExtraCondition:=ConveyorIO70159.xEmpty AND NOT ConveyorIO70159.xCWPresent AND NOT ConveyorIO701102.xCWPresent;
(*
ComConveyorIO70159.i_iResponsPCPLC:=D2540; 
ComConveyorIO70159.i_iTypeInfoPCPLC:=D2541;
ComConveyorIO70159.i_iReadWriteFlagPCPLC:=D2545; 
ComConveyorIO70159.i_iTaskProcessFlagPCPLC:=D2546; 
ComConveyorIO70159.i_iCommandPCPLC:=D2547; 
ComConveyorIO70159.i_iTaskIDPCPLC:=D2548; 
DMOV(TRUE,D2549,ComConveyorIO70159.i_diDestinationDevicePCPLC); 
ComConveyorIO70159.i_iProductIDPCPLC:=D2551;
D3540:=ComConveyorIO70159.o_iRequestPLCPC; 
D3541:=ComConveyorIO70159.o_iForceInportPLCPC;
D3542:=ComConveyorIO70159.o_iFolderNumberPLCPC;
D3543:=ComConveyorIO70159.o_iEmptyPLCPC;
D3545:=ComConveyorIO70159.o_iReadWriteFlagPLCPC; 
D3546:=ComConveyorIO70159.o_iDeviceStatusPLCPC; 
D3547:=ComConveyorIO70159.o_iTaskIDPLCPC; 
D3548:=ComConveyorIO70159.o_iProductIDPLCPC;
ComConveyorIO70159.i_xExportConveyor:=1;
*)
ComConveyorIO701120.i_iResponsPCPLC:=D2555; 
ComConveyorIO701120.i_iTypeInfoPCPLC:=D2556;
ComConveyorIO701120.i_iReadWriteFlagPCPLC:=D2560; 
ComConveyorIO701120.i_iTaskProcessFlagPCPLC:=D2561; 
ComConveyorIO701120.i_iCommandPCPLC:=D2562; 
ComConveyorIO701120.i_iTaskIDPCPLC:=D2563; 
DMOV(TRUE,D2564,ComConveyorIO701120.i_diDestinationDevicePCPLC); 
ComConveyorIO701120.i_iProductIDPCPLC:=D2566;
D3555:=ComConveyorIO701120.o_iRequestPLCPC; 
D3556:=ComConveyorIO701120.o_iForceInportPLCPC;
D3557:=ComConveyorIO701120.o_iFolderNumberPLCPC;
D3558:=ComConveyorIO701120.o_iEmptyPLCPC;
D3560:=ComConveyorIO701120.o_iReadWriteFlagPLCPC; 
D3561:=ComConveyorIO701120.o_iDeviceStatusPLCPC; 
D3562:=ComConveyorIO701120.o_iTaskIDPLCPC; 
D3563:=ComConveyorIO701120.o_iProductIDPLCPC;
ComConveyorIO701120.i_xExportConveyor:=1;
ComConveyorIO701120.i_xExtraCondition:=ConveyorIO701119.xEmpty AND NOT ConveyorIO701119.xCWPresent AND NOT ConveyorIO701120.xCWPresent;
(*
ComConveyorIO701119.i_iResponsPCPLC:=D2570; 
ComConveyorIO701119.i_iTypeInfoPCPLC:=D2571;
ComConveyorIO701119.i_iReadWriteFlagPCPLC:=D2575; 
ComConveyorIO701119.i_iTaskProcessFlagPCPLC:=D2576; 
ComConveyorIO701119.i_iCommandPCPLC:=D2577; 
ComConveyorIO701119.i_iTaskIDPCPLC:=D2578; 
DMOV(TRUE,D2579,ComConveyorIO701119.i_diDestinationDevicePCPLC); 
ComConveyorIO701119.i_iProductIDPCPLC:=D2581;
D3570:=ComConveyorIO701119.o_iRequestPLCPC; 
D3571:=ComConveyorIO701119.o_iForceInportPLCPC;
D3572:=ComConveyorIO701119.o_iFolderNumberPLCPC;
D3573:=ComConveyorIO701119.o_iEmptyPLCPC;
D3575:=ComConveyorIO701119.o_iReadWriteFlagPLCPC; 
D3576:=ComConveyorIO701119.o_iDeviceStatusPLCPC; 
D3577:=ComConveyorIO701119.o_iTaskIDPLCPC; 
D3578:=ComConveyorIO701119.o_iProductIDPLCPC;
ComConveyorIO701119.i_xExportConveyor:=1;*)